(* CODESYS project CodeSys_main_v2.project (continued)
  5ce3da45-db07-42e7-a21c-a00fff4ed8f6|C:\Users\ggb\Documents\#PROJECTS\2016_06_29_Denmark\Visu\CheckBox_1.png
  5ce3da45-db07-42e7-a21c-a00fff4ed8f6|C:\Users\ggb\Documents\#PROJECTS\2016_06_29_Denmark\Visu\Manual_1.png
  5ce3da45-db07-42e7-a21c-a00fff4ed8f6|C:\Users\ggb\Documents\#PROJECTS\2016_06_29_Denmark\Pictures\071-030_Modul Trocknen.jpg
  5ce3da45-db07-42e7-a21c-a00fff4ed8f6|C:\Users\ggb\Documents\#PROJECTS\2016_06_29_Denmark\Visu\English.gif
  5ce3da45-db07-42e7-a21c-a00fff4ed8f6|C:\Users\ggb\Documents\#PROJECTS\2016_06_29_Denmark\Visu\Home_1.png
  5ce3da45-db07-42e7-a21c-a00fff4ed8f6|C:\Users\ggb\Documents\#PROJECTS\2016_06_29_Denmark\Visu\LeftArrow_Bold.png
  5ce3da45-db07-42e7-a21c-a00fff4ed8f6|C:\Users\ggb\Documents\#PROJECTS\2016_06_29_Denmark\Pictures\071-050a_Bohren EA.jpg
  5ce3da45-db07-42e7-a21c-a00fff4ed8f6|C:\Users\ggb\Documents\#PROJECTS\2016_06_29_Denmark\Visu\Parameters_0.png
  Data Types/
    HMI and SCADA/
      data type st_WinCC
      data type st_ManualWorkplace
      CDPX/
        data type st_StopperSensorSignals
        data type st_InterctiveErrors
        data type st_Errors
        data type st_ConveyorSignals
        data type st_AppButtonControl
        data type st_StopperButtonState
        data type st_CdpxButtonState
        data type st_AppSensors
        data type st_ConveyorButtonState
      data type st_ButtonState
      data type st_TransitionData
    SAP/
      sub_structures/
        data type st_Par_Req
        data type st_Start_Req
        data type st_Com
        data type st_Start_Res
        data type st_Comp_Req
        data type st_Comp_Res
      ManualWork/
        data type st_MesRcvData_ManualWork
      data type st_CompleteSfc
      data type st_ParametricData
      data type st_StartSfc
    Error/
      data type st_InteractiveError
      data type st_RobotError
      data type u_Error
      data type st_Error
      data type st_ErrorWords
      data type st_ErrorEvent
    data type st_GetShuntId
    Application/
      data type st_AppControl
      data type st_AppSettings
      data type st_AppState
      data type st_AppInfo
  5ce3da45-db07-42e7-a21c-a00fff4ed8f6|C:\Users\ggb\Documents\#PROJECTS\2016_06_29_Denmark\Visu\Plus.png
  5ce3da45-db07-42e7-a21c-a00fff4ed8f6|C:\Users\ggb\Documents\#PROJECTS\2016_06_29_Denmark\Visu\Settings_1.png
  5ce3da45-db07-42e7-a21c-a00fff4ed8f6|C:\Users\ggb\Documents\#PROJECTS\2016_06_29_Denmark\Visu\Settings_0.png
  5ce3da45-db07-42e7-a21c-a00fff4ed8f6|C:\Users\ggb\Documents\#PROJECTS\2016_06_29_Denmark\Visu\Settings_0.png
  5ce3da45-db07-42e7-a21c-a00fff4ed8f6|C:\Users\ggb\Documents\#PROJECTS\2016_06_29_Denmark\Visu\Parameters_1.png
  5ce3da45-db07-42e7-a21c-a00fff4ed8f6|C:\Users\ggb\Documents\#PROJECTS\2016_06_29_Denmark\Visu\English.gif
  5ce3da45-db07-42e7-a21c-a00fff4ed8f6|C:\Users\ggb\Documents\#PROJECTS\2016_06_29_Denmark\Visu\RightArrow.png
  5ce3da45-db07-42e7-a21c-a00fff4ed8f6|C:\Users\ggb\Documents\#PROJECTS\2016_06_29_Denmark\Pictures\071-050a_Bohren EA.jpg
  5ce3da45-db07-42e7-a21c-a00fff4ed8f6|C:\Users\ggb\Documents\#PROJECTS\2016_06_29_Denmark\Visu\CheckBox_0.png
  5ce3da45-db07-42e7-a21c-a00fff4ed8f6|C:\Users\ggb\Documents\#PROJECTS\2016_06_29_Denmark\Visu\English.gif
  5ce3da45-db07-42e7-a21c-a00fff4ed8f6|C:\Users\ggb\Documents\#PROJECTS\2016_06_29_Denmark\Visu\Stopper.jpg
  5ce3da45-db07-42e7-a21c-a00fff4ed8f6|C:\Users\ggb\Documents\#PROJECTS\2016_06_29_Denmark\Visu\CheckBox_1.png
  5ce3da45-db07-42e7-a21c-a00fff4ed8f6|C:\Users\ggb\Documents\#PROJECTS\2016_06_29_Denmark\Visu\Plus.png
  5ce3da45-db07-42e7-a21c-a00fff4ed8f6|C:\Users\ggb\Documents\#PROJECTS\2016_06_29_Denmark\Pictures\071-046b_Magazin.jpg
  5ce3da45-db07-42e7-a21c-a00fff4ed8f6|C:\Users\ggb\Documents\#PROJECTS\2016_06_29_Denmark\Pictures\cpFactory_Conveyor.png
  5ce3da45-db07-42e7-a21c-a00fff4ed8f6|C:\Users\ggb\Documents\#PROJECTS\2016_06_29_Denmark\Visu\English.gif
  5ce3da45-db07-42e7-a21c-a00fff4ed8f6|C:\Users\ggb\Documents\#PROJECTS\2016_06_29_Denmark\Visu\Parameters_1.png
  5ce3da45-db07-42e7-a21c-a00fff4ed8f6|C:\Users\ggb\Documents\#PROJECTS\2016_06_29_Denmark\Visu\RightArrow.png
  5ce3da45-db07-42e7-a21c-a00fff4ed8f6|C:\Users\ggb\Documents\#PROJECTS\2016_06_29_Denmark\Visu\LeftArrow_Bold.png
  5ce3da45-db07-42e7-a21c-a00fff4ed8f6|C:\Users\ggb\Documents\#PROJECTS\2016_06_29_Denmark\Visu\Manual_1.png
  5ce3da45-db07-42e7-a21c-a00fff4ed8f6|C:\Users\ggb\Documents\#PROJECTS\2016_06_29_Denmark\Visu\Plus.png
  5ce3da45-db07-42e7-a21c-a00fff4ed8f6|C:\Users\ggb\Documents\#PROJECTS\2016_06_29_Denmark\Visu\FESTO.png
  5ce3da45-db07-42e7-a21c-a00fff4ed8f6|C:\Users\ggb\Documents\#PROJECTS\2016_06_29_Denmark\Visu\Parameters_0.png
  5ce3da45-db07-42e7-a21c-a00fff4ed8f6|C:\Users\ggb\Documents\#PROJECTS\2016_06_29_Denmark\Pictures\071-046b_Magazin.jpg
  5ce3da45-db07-42e7-a21c-a00fff4ed8f6|C:\Users\ggb\Documents\#PROJECTS\2016_06_29_Denmark\Visu\LeftArrow_Bold.png
  5ce3da45-db07-42e7-a21c-a00fff4ed8f6|C:\Users\ggb\Documents\#PROJECTS\2016_06_29_Denmark\Visu\Home_0.png
  5ce3da45-db07-42e7-a21c-a00fff4ed8f6|C:\Users\ggb\Documents\#PROJECTS\2016_06_29_Denmark\Visu\Home_1.png
  5ce3da45-db07-42e7-a21c-a00fff4ed8f6|C:\Users\ggb\Documents\#PROJECTS\2016_06_29_Denmark\Visu\German.gif
  5ce3da45-db07-42e7-a21c-a00fff4ed8f6|C:\Users\ggb\Documents\#PROJECTS\2016_06_29_Denmark\Visu\Stopper.jpg
  5ce3da45-db07-42e7-a21c-a00fff4ed8f6|C:\Users\ggb\Documents\#PROJECTS\2016_06_29_Denmark\Visu\RightArrow.png
  5ce3da45-db07-42e7-a21c-a00fff4ed8f6|C:\Users\ggb\Documents\#PROJECTS\2016_06_29_Denmark\Visu\Home_0.png
  5ce3da45-db07-42e7-a21c-a00fff4ed8f6|C:\Users\ggb\Documents\#PROJECTS\2016_06_29_Denmark\Visu\Home_1.png
  5ce3da45-db07-42e7-a21c-a00fff4ed8f6|C:\Users\ggb\Documents\#PROJECTS\2016_06_29_Denmark\Visu\Home_1.png
  5ce3da45-db07-42e7-a21c-a00fff4ed8f6|C:\Users\ggb\Documents\#PROJECTS\2016_06_29_Denmark\Visu\FESTO.png
  5ce3da45-db07-42e7-a21c-a00fff4ed8f6|C:\Users\ggb\Documents\#PROJECTS\2016_06_29_Denmark\Visu\Home_1.png
  5ce3da45-db07-42e7-a21c-a00fff4ed8f6|C:\Users\ggb\Documents\#PROJECTS\2016_06_29_Denmark\Visu\CheckBox_1.png
  5ce3da45-db07-42e7-a21c-a00fff4ed8f6|C:\Users\ggb\Documents\#PROJECTS\2016_06_29_Denmark\Visu\CheckBox_0.png
  5ce3da45-db07-42e7-a21c-a00fff4ed8f6|C:\Users\ggb\Documents\#PROJECTS\2016_06_29_Denmark\Visu\CheckBox_0.png
  5ce3da45-db07-42e7-a21c-a00fff4ed8f6|C:\Users\ggb\Documents\#PROJECTS\2016_06_29_Denmark\Pictures\Cam.jpg
  5ce3da45-db07-42e7-a21c-a00fff4ed8f6|C:\Users\ggb\Documents\#PROJECTS\2016_06_29_Denmark\Visu\Settings_1.png
  5ce3da45-db07-42e7-a21c-a00fff4ed8f6|C:\Users\ggb\Documents\#PROJECTS\2016_06_29_Denmark\Visu\RightArrow_Bold.png
  5ce3da45-db07-42e7-a21c-a00fff4ed8f6|C:\Users\ggb\Documents\#PROJECTS\2016_06_29_Denmark\Visu\RightArrow_Bold.png
  5ce3da45-db07-42e7-a21c-a00fff4ed8f6|C:\Users\ggb\Documents\#PROJECTS\2016_06_29_Denmark\Visu\CheckBox_1.png
  5ce3da45-db07-42e7-a21c-a00fff4ed8f6|C:\Users\ggb\Documents\#PROJECTS\2016_06_29_Denmark\Visu\Settings_0.png
  5ce3da45-db07-42e7-a21c-a00fff4ed8f6|C:\Users\ggb\Documents\#PROJECTS\2016_06_29_Denmark\Visu\Home_0.png
  5ce3da45-db07-42e7-a21c-a00fff4ed8f6|C:\Users\ggb\Documents\#PROJECTS\2016_06_29_Denmark\Pictures\cpFactory_Bypass.png
  5ce3da45-db07-42e7-a21c-a00fff4ed8f6|C:\Users\ggb\Documents\#PROJECTS\2016_06_29_Denmark\Visu\LeftArrow_Bold.png
  5ce3da45-db07-42e7-a21c-a00fff4ed8f6|C:\Users\ggb\Documents\#PROJECTS\2016_06_29_Denmark\Visu\RightArrow.png
  5ce3da45-db07-42e7-a21c-a00fff4ed8f6|C:\Users\ggb\Documents\#PROJECTS\2016_06_29_Denmark\Visu\RightArrow.png
  5ce3da45-db07-42e7-a21c-a00fff4ed8f6|C:\Users\ggb\Documents\#PROJECTS\2016_06_29_Denmark\Visu\RightArrow_Bold.png
  5ce3da45-db07-42e7-a21c-a00fff4ed8f6|C:\Users\ggb\Documents\#PROJECTS\2016_06_29_Denmark\Visu\FESTO.png
  5ce3da45-db07-42e7-a21c-a00fff4ed8f6|C:\Users\ggb\Documents\#PROJECTS\2016_06_29_Denmark\Pictures\cpFactory_Bypass.png
  5ce3da45-db07-42e7-a21c-a00fff4ed8f6|C:\Users\ggb\Documents\#PROJECTS\2016_06_29_Denmark\Visu\Settings_0.png
  5ce3da45-db07-42e7-a21c-a00fff4ed8f6|C:\Users\ggb\Documents\#PROJECTS\2016_06_29_Denmark\Pictures\071-030_Modul Trocknen.jpg
  5ce3da45-db07-42e7-a21c-a00fff4ed8f6|C:\Users\ggb\Documents\#PROJECTS\2016_06_29_Denmark\Visu\RightArrow_Bold.png
  5ce3da45-db07-42e7-a21c-a00fff4ed8f6|C:\Users\ggb\Documents\#PROJECTS\2016_06_29_Denmark\Pictures\071-046b_Magazin.jpg
  5ce3da45-db07-42e7-a21c-a00fff4ed8f6|C:\Users\ggb\Documents\#PROJECTS\2016_06_29_Denmark\Pictures\cpFactory_Bypass.png
  Programs/
    function block TrafficStopper [ST]: _DefaultMode, _ModuleCalls
    function block StopperWithMes [ST]: _MesMode, _DefaultMode, _ModuleCalls, _SapMode
    function block SwitchWithoutMes [ST]: _SapMode, _MesMode, _DefaultMode, _ModuleCalls
    Tools/
      function block ErrorFifo [ST]
      function block MovCntr2B2M [LD]
      function DateFormat [ST]
      function block MovCntr3B3M [LD]
      program ErrorCpyHMI [ST]
      program ErrorCpyWinCC [ST]
    Visu/
      program VisuProgramStp [ST]
    function block SwitchWithMes [ST]: _DefaultMode, _ModuleCalls, _SapMode, _MesMode
  5ce3da45-db07-42e7-a21c-a00fff4ed8f6|C:\Users\ggb\Documents\#PROJECTS\2016_06_29_Denmark\Visu\Home_1.png
  5ce3da45-db07-42e7-a21c-a00fff4ed8f6|C:\Users\ggb\Documents\#PROJECTS\2016_06_29_Denmark\Pictures\cpFactory_Bypass.png
  5ce3da45-db07-42e7-a21c-a00fff4ed8f6|C:\Users\ggb\Documents\#PROJECTS\2016_06_29_Denmark\Visu\CheckBox_0.png
  5ce3da45-db07-42e7-a21c-a00fff4ed8f6|C:\Users\ggb\Documents\#PROJECTS\2016_06_29_Denmark\Pictures\071-046b_Magazin.jpg
  5ce3da45-db07-42e7-a21c-a00fff4ed8f6|C:\Users\ggb\Documents\#PROJECTS\2016_06_29_Denmark\Visu\German.gif
  5ce3da45-db07-42e7-a21c-a00fff4ed8f6|C:\Users\ggb\Documents\#PROJECTS\2016_06_29_Denmark\Visu\RightArrow_Bold.png
  5ce3da45-db07-42e7-a21c-a00fff4ed8f6|C:\Users\ggb\Documents\#PROJECTS\2016_06_29_Denmark\Visu\English.gif
  5ce3da45-db07-42e7-a21c-a00fff4ed8f6|C:\Users\ggb\Documents\#PROJECTS\2016_06_29_Denmark\Pictures\Kuka_Agilus.png
  5ce3da45-db07-42e7-a21c-a00fff4ed8f6|C:\Users\ggb\Documents\#PROJECTS\2016_06_29_Denmark\Visu\Parameters_1.png
  5ce3da45-db07-42e7-a21c-a00fff4ed8f6|C:\Users\ggb\Documents\#PROJECTS\2016_06_29_Denmark\Visu\FESTO.png
  5ce3da45-db07-42e7-a21c-a00fff4ed8f6|C:\Users\ggb\Documents\#PROJECTS\2016_06_29_Denmark\Pictures\071-046b_Magazin.jpg
  5ce3da45-db07-42e7-a21c-a00fff4ed8f6|C:\Users\ggb\Documents\#PROJECTS\2016_06_29_Denmark\Visu\German.gif
  5ce3da45-db07-42e7-a21c-a00fff4ed8f6|C:\Users\ggb\Documents\#PROJECTS\2016_06_29_Denmark\Visu\Settings_0.png
  5ce3da45-db07-42e7-a21c-a00fff4ed8f6|C:\Users\ggb\Documents\#PROJECTS\2016_06_29_Denmark\Visu\Plus.png
  5ce3da45-db07-42e7-a21c-a00fff4ed8f6|C:\Users\ggb\Documents\#PROJECTS\2016_06_29_Denmark\Visu\Settings_1.png
  5ce3da45-db07-42e7-a21c-a00fff4ed8f6|C:\Users\ggb\Documents\#PROJECTS\2016_06_29_Denmark\Visu\Settings_0.png
  5ce3da45-db07-42e7-a21c-a00fff4ed8f6|C:\Users\ggb\Documents\#PROJECTS\2016_06_29_Denmark\Visu\CheckBox_1.png
  5ce3da45-db07-42e7-a21c-a00fff4ed8f6|C:\Users\ggb\Documents\#PROJECTS\2016_06_29_Denmark\Visu\German.gif
  5ce3da45-db07-42e7-a21c-a00fff4ed8f6|C:\Users\ggb\Documents\#PROJECTS\2016_06_29_Denmark\Visu\Plus.png
  5ce3da45-db07-42e7-a21c-a00fff4ed8f6|C:\Users\ggb\Documents\#PROJECTS\2016_06_29_Denmark\Pictures\071-060_Kameraprüfen.jpg
  5ce3da45-db07-42e7-a21c-a00fff4ed8f6|C:\Users\ggb\Documents\#PROJECTS\2016_06_29_Denmark\Visu\Manual_0.png
  5ce3da45-db07-42e7-a21c-a00fff4ed8f6|C:\Users\ggb\Documents\#PROJECTS\2016_06_29_Denmark\Visu\Settings_1.png
  5ce3da45-db07-42e7-a21c-a00fff4ed8f6|C:\Users\ggb\Documents\#PROJECTS\2016_06_29_Denmark\Pictures\071-050a_Bohren EA.jpg
  5ce3da45-db07-42e7-a21c-a00fff4ed8f6|C:\Users\ggb\Documents\#PROJECTS\2016_06_29_Denmark\Visu\Settings_1.png
  5ce3da45-db07-42e7-a21c-a00fff4ed8f6|C:\Users\ggb\Documents\#PROJECTS\2016_06_29_Denmark\Pictures\071-030_Modul Trocknen.jpg
  5ce3da45-db07-42e7-a21c-a00fff4ed8f6|C:\Users\ggb\Documents\#PROJECTS\2016_06_29_Denmark\Visu\LeftArrow_Bold.png
  5ce3da45-db07-42e7-a21c-a00fff4ed8f6|C:\Users\ggb\Documents\#PROJECTS\2016_06_29_Denmark\Pictures\071-030_Modul Trocknen.jpg
  5ce3da45-db07-42e7-a21c-a00fff4ed8f6|C:\Users\ggb\Documents\#PROJECTS\2016_06_29_Denmark\Pictures\071-046b_Magazin.jpg
  5ce3da45-db07-42e7-a21c-a00fff4ed8f6|C:\Users\ggb\Documents\#PROJECTS\2016_06_29_Denmark\Pictures\cpFactory_Bypass.png
  5ce3da45-db07-42e7-a21c-a00fff4ed8f6|C:\Users\ggb\Documents\#PROJECTS\2016_06_29_Denmark\Visu\Plus.png
  5ce3da45-db07-42e7-a21c-a00fff4ed8f6|C:\Users\ggb\Documents\#PROJECTS\2016_06_29_Denmark\Visu\FESTO.png
  5ce3da45-db07-42e7-a21c-a00fff4ed8f6|C:\Users\ggb\Documents\#PROJECTS\2016_06_29_Denmark\Visu\English.gif
  5ce3da45-db07-42e7-a21c-a00fff4ed8f6|C:\Users\ggb\Documents\#PROJECTS\2016_06_29_Denmark\Visu\Stopper.jpg
  5ce3da45-db07-42e7-a21c-a00fff4ed8f6|C:\Users\ggb\Documents\#PROJECTS\2016_06_29_Denmark\Visu\Stopper.jpg
  5ce3da45-db07-42e7-a21c-a00fff4ed8f6|C:\Users\ggb\Documents\#PROJECTS\2016_06_29_Denmark\Pictures\071-030_Modul Trocknen.jpg
  5ce3da45-db07-42e7-a21c-a00fff4ed8f6|C:\Users\ggb\Documents\#PROJECTS\2016_06_29_Denmark\Pictures\cpFactory_Bypass.png
  5ce3da45-db07-42e7-a21c-a00fff4ed8f6|C:\Users\ggb\Documents\#PROJECTS\2016_06_29_Denmark\Visu\CheckBox_0.png
  5ce3da45-db07-42e7-a21c-a00fff4ed8f6|C:\Users\ggb\Documents\#PROJECTS\2016_06_29_Denmark\Visu\CheckBox_0.png
  5ce3da45-db07-42e7-a21c-a00fff4ed8f6|C:\Users\ggb\Documents\#PROJECTS\2016_06_29_Denmark\Visu\Stopper.jpg
  5ce3da45-db07-42e7-a21c-a00fff4ed8f6|C:\Users\ggb\Documents\#PROJECTS\2016_06_29_Denmark\Pictures\cpFactory_Conveyor.png
  5ce3da45-db07-42e7-a21c-a00fff4ed8f6|C:\Users\ggb\Documents\#PROJECTS\2016_06_29_Denmark\Visu\Settings_0.png
  5ce3da45-db07-42e7-a21c-a00fff4ed8f6|C:\Users\ggb\Documents\#PROJECTS\2016_06_29_Denmark\Visu\Parameters_0.png
  5ce3da45-db07-42e7-a21c-a00fff4ed8f6|C:\Users\ggb\Documents\#PROJECTS\2016_06_29_Denmark\Visu\Home_1.png
  5ce3da45-db07-42e7-a21c-a00fff4ed8f6|C:\Users\ggb\Documents\#PROJECTS\2016_06_29_Denmark\Pictures\071-050a_Bohren EA.jpg
  5ce3da45-db07-42e7-a21c-a00fff4ed8f6|C:\Users\ggb\Documents\#PROJECTS\2016_06_29_Denmark\Visu\Manual_1.png
  5ce3da45-db07-42e7-a21c-a00fff4ed8f6|C:\Users\ggb\Documents\#PROJECTS\2016_06_29_Denmark\Visu\Stopper.jpg
  5ce3da45-db07-42e7-a21c-a00fff4ed8f6|C:\Users\ggb\Documents\#PROJECTS\2016_06_29_Denmark\Pictures\071-030_Modul Trocknen.jpg
  5ce3da45-db07-42e7-a21c-a00fff4ed8f6|C:\Users\ggb\Documents\#PROJECTS\2016_06_29_Denmark\Visu\CheckBox_0.png
  5ce3da45-db07-42e7-a21c-a00fff4ed8f6|C:\Users\ggb\Documents\#PROJECTS\2016_06_29_Denmark\Visu\CheckBox_1.png
  5ce3da45-db07-42e7-a21c-a00fff4ed8f6|C:\Users\ggb\Documents\#PROJECTS\2016_06_29_Denmark\Visu\LeftArrow_Bold.png
  5ce3da45-db07-42e7-a21c-a00fff4ed8f6|C:\Users\ggb\Documents\#PROJECTS\2016_06_29_Denmark\Pictures\cpFactory_Bypass.png
  5ce3da45-db07-42e7-a21c-a00fff4ed8f6|C:\Users\ggb\Documents\#PROJECTS\2016_06_29_Denmark\Visu\LeftArrow_Bold.png
  Global Variables/
    global variables fromCDPX
    global variables Standards
    global variables toCDPX
    global variables SAP
    global variables SAPInit
    global variables SAPHMI
  5ce3da45-db07-42e7-a21c-a00fff4ed8f6|C:\Users\ggb\Documents\#PROJECTS\2016_06_29_Denmark\Visu\CheckBox_0.png
  5ce3da45-db07-42e7-a21c-a00fff4ed8f6|C:\Users\ggb\Documents\#PROJECTS\2016_06_29_Denmark\Pictures\cpFactory_Conveyor.png
  5ce3da45-db07-42e7-a21c-a00fff4ed8f6|C:\Users\ggb\Documents\#PROJECTS\2016_06_29_Denmark\Pictures\071-046b_Magazin.jpg
  5ce3da45-db07-42e7-a21c-a00fff4ed8f6|C:\Users\ggb\Documents\#PROJECTS\2016_06_29_Denmark\Visu\RightArrow.png
  5ce3da45-db07-42e7-a21c-a00fff4ed8f6|C:\Users\ggb\Documents\#PROJECTS\2016_06_29_Denmark\Pictures\cpFactory_Bypass.png
  5ce3da45-db07-42e7-a21c-a00fff4ed8f6|C:\Users\ggb\Documents\#PROJECTS\2016_06_29_Denmark\Pictures\071-060_Kameraprüfen.jpg
  5ce3da45-db07-42e7-a21c-a00fff4ed8f6|C:\Users\ggb\Documents\#PROJECTS\2016_06_29_Denmark\Visu\German.gif
  5ce3da45-db07-42e7-a21c-a00fff4ed8f6|C:\Users\ggb\Documents\#PROJECTS\2016_06_29_Denmark\Visu\CheckBox_0.png
  5ce3da45-db07-42e7-a21c-a00fff4ed8f6|C:\Users\ggb\Documents\#PROJECTS\2016_06_29_Denmark\Visu\Settings_0.png
  5ce3da45-db07-42e7-a21c-a00fff4ed8f6|C:\Users\ggb\Documents\#PROJECTS\2016_06_29_Denmark\Visu\CheckBox_1.png
  5ce3da45-db07-42e7-a21c-a00fff4ed8f6|C:\Users\ggb\Documents\#PROJECTS\2016_06_29_Denmark\Visu\FESTO.png
  5ce3da45-db07-42e7-a21c-a00fff4ed8f6|C:\Users\ggb\Documents\#PROJECTS\2016_06_29_Denmark\Visu\CheckBox_0.png
  5ce3da45-db07-42e7-a21c-a00fff4ed8f6|C:\Users\ggb\Documents\#PROJECTS\2016_06_29_Denmark\Pictures\cpFactory_Conveyor.png
  5ce3da45-db07-42e7-a21c-a00fff4ed8f6|C:\Users\ggb\Documents\#PROJECTS\2016_06_29_Denmark\Visu\CheckBox_1.png
  5ce3da45-db07-42e7-a21c-a00fff4ed8f6|C:\Users\ggb\Documents\#PROJECTS\2016_06_29_Denmark\Pictures\cpFactory_Conveyor.png
  5ce3da45-db07-42e7-a21c-a00fff4ed8f6|C:\Users\ggb\Documents\#PROJECTS\2016_06_29_Denmark\Pictures\071-050a_Bohren EA.jpg
  5ce3da45-db07-42e7-a21c-a00fff4ed8f6|C:\Users\ggb\Documents\#PROJECTS\2016_06_29_Denmark\Visu\Parameters_0.png
  5ce3da45-db07-42e7-a21c-a00fff4ed8f6|C:\Users\ggb\Documents\#PROJECTS\2016_06_29_Denmark\Visu\CheckBox_1.png
  5ce3da45-db07-42e7-a21c-a00fff4ed8f6|C:\Users\ggb\Documents\#PROJECTS\2016_06_29_Denmark\Visu\Home_1.png
  5ce3da45-db07-42e7-a21c-a00fff4ed8f6|C:\Users\ggb\Documents\#PROJECTS\2016_06_29_Denmark\Pictures\071-060_Kameraprüfen.jpg
  5ce3da45-db07-42e7-a21c-a00fff4ed8f6|C:\Users\ggb\Documents\#PROJECTS\2016_06_29_Denmark\Visu\English.gif
  5ce3da45-db07-42e7-a21c-a00fff4ed8f6|C:\Users\ggb\Documents\#PROJECTS\2016_06_29_Denmark\Pictures\cpFactory_Bypass.png
  5ce3da45-db07-42e7-a21c-a00fff4ed8f6|C:\Users\ggb\Documents\#PROJECTS\2016_06_29_Denmark\Visu\Parameters_1.png
  5ce3da45-db07-42e7-a21c-a00fff4ed8f6|C:\Users\ggb\Documents\#PROJECTS\2016_06_29_Denmark\Visu\Manual_1.png
  5ce3da45-db07-42e7-a21c-a00fff4ed8f6|C:\Users\ggb\Documents\#PROJECTS\2016_06_29_Denmark\Visu\CheckBox_0.png
  5ce3da45-db07-42e7-a21c-a00fff4ed8f6|C:\Users\ggb\Documents\#PROJECTS\2016_06_29_Denmark\Visu\Manual_0.png
  5ce3da45-db07-42e7-a21c-a00fff4ed8f6|C:\Users\ggb\Documents\#PROJECTS\2016_06_29_Denmark\Visu\Manual_0.png
  5ce3da45-db07-42e7-a21c-a00fff4ed8f6|C:\Users\ggb\Documents\#PROJECTS\2016_06_29_Denmark\Visu\Home_1.png
  5ce3da45-db07-42e7-a21c-a00fff4ed8f6|C:\Users\ggb\Documents\#PROJECTS\2016_06_29_Denmark\Pictures\071-046b_Magazin.jpg
  5ce3da45-db07-42e7-a21c-a00fff4ed8f6|C:\Users\ggb\Documents\#PROJECTS\2016_06_29_Denmark\Visu\English.gif
  5ce3da45-db07-42e7-a21c-a00fff4ed8f6|C:\Users\ggb\Documents\#PROJECTS\2016_06_29_Denmark\Pictures\cpFactory_Conveyor.png
  5ce3da45-db07-42e7-a21c-a00fff4ed8f6|C:\Users\ggb\Documents\#PROJECTS\2016_06_29_Denmark\Pictures\071-050a_Bohren EA.jpg
  5ce3da45-db07-42e7-a21c-a00fff4ed8f6|C:\Users\ggb\Documents\#PROJECTS\2016_06_29_Denmark\Visu\English.gif
  5ce3da45-db07-42e7-a21c-a00fff4ed8f6|C:\Users\ggb\Documents\#PROJECTS\2016_06_29_Denmark\Visu\Parameters_1.png
  5ce3da45-db07-42e7-a21c-a00fff4ed8f6|C:\Users\ggb\Documents\#PROJECTS\2016_06_29_Denmark\Visu\RightArrow_Bold.png
  5ce3da45-db07-42e7-a21c-a00fff4ed8f6|C:\Users\ggb\Documents\#PROJECTS\2016_06_29_Denmark\Visu\FESTO.png
  5ce3da45-db07-42e7-a21c-a00fff4ed8f6|C:\Users\ggb\Documents\#PROJECTS\2016_06_29_Denmark\Pictures\071-050a_Bohren EA.jpg
  5ce3da45-db07-42e7-a21c-a00fff4ed8f6|C:\Users\ggb\Documents\#PROJECTS\2016_06_29_Denmark\Pictures\071-046b_Magazin.jpg
  5ce3da45-db07-42e7-a21c-a00fff4ed8f6|C:\Users\ggb\Documents\#PROJECTS\2016_06_29_Denmark\Visu\RightArrow_Bold.png
  5ce3da45-db07-42e7-a21c-a00fff4ed8f6|C:\Users\ggb\Documents\#PROJECTS\2016_06_29_Denmark\Visu\Parameters_0.png
  5ce3da45-db07-42e7-a21c-a00fff4ed8f6|C:\Users\ggb\Documents\#PROJECTS\2016_06_29_Denmark\Pictures\cpFactory_Conveyor.png
  5ce3da45-db07-42e7-a21c-a00fff4ed8f6|C:\Users\ggb\Documents\#PROJECTS\2016_06_29_Denmark\Visu\Home_0.png
  5ce3da45-db07-42e7-a21c-a00fff4ed8f6|C:\Users\ggb\Documents\#PROJECTS\2016_06_29_Denmark\Visu\LeftArrow_Bold.png
  5ce3da45-db07-42e7-a21c-a00fff4ed8f6|C:\Users\ggb\Documents\#PROJECTS\2016_06_29_Denmark\Visu\Parameters_0.png
  5ce3da45-db07-42e7-a21c-a00fff4ed8f6|C:\Users\ggb\Documents\#PROJECTS\2016_06_29_Denmark\Visu\Manual_0.png
  5ce3da45-db07-42e7-a21c-a00fff4ed8f6|C:\Users\ggb\Documents\#PROJECTS\2016_06_29_Denmark\Visu\Manual_0.png
  5ce3da45-db07-42e7-a21c-a00fff4ed8f6|C:\Users\ggb\Documents\#PROJECTS\2016_06_29_Denmark\Visu\Settings_1.png
  5ce3da45-db07-42e7-a21c-a00fff4ed8f6|C:\Users\ggb\Documents\#PROJECTS\2016_06_29_Denmark\Visu\Home_0.png
  5ce3da45-db07-42e7-a21c-a00fff4ed8f6|C:\Users\ggb\Documents\#PROJECTS\2016_06_29_Denmark\Visu\FESTO.png
  5ce3da45-db07-42e7-a21c-a00fff4ed8f6|C:\Users\ggb\Documents\#PROJECTS\2016_06_29_Denmark\Visu\German.gif
  5ce3da45-db07-42e7-a21c-a00fff4ed8f6|C:\Users\ggb\Documents\#PROJECTS\2016_06_29_Denmark\Visu\Settings_0.png
  5ce3da45-db07-42e7-a21c-a00fff4ed8f6|C:\Users\ggb\Documents\#PROJECTS\2016_06_29_Denmark\Visu\RightArrow_Bold.png
  5ce3da45-db07-42e7-a21c-a00fff4ed8f6|C:\Users\ggb\Documents\#PROJECTS\2016_06_29_Denmark\Visu\Stopper.jpg
  5ce3da45-db07-42e7-a21c-a00fff4ed8f6|C:\Users\ggb\Documents\#PROJECTS\2016_06_29_Denmark\Visu\Parameters_1.png
  5ce3da45-db07-42e7-a21c-a00fff4ed8f6|C:\Users\ggb\Documents\#PROJECTS\2016_06_29_Denmark\Visu\FESTO.png
  5ce3da45-db07-42e7-a21c-a00fff4ed8f6|C:\Users\ggb\Documents\#PROJECTS\2016_06_29_Denmark\Visu\German.gif
  5ce3da45-db07-42e7-a21c-a00fff4ed8f6|C:\Users\ggb\Documents\#PROJECTS\2016_06_29_Denmark\Visu\Home_0.png
  text list GlobalTextList
  5ce3da45-db07-42e7-a21c-a00fff4ed8f6|C:\Users\ggb\Documents\#PROJECTS\2016_06_29_Denmark\Visu\FESTO.png
  5ce3da45-db07-42e7-a21c-a00fff4ed8f6|C:\Users\ggb\Documents\#PROJECTS\2016_06_29_Denmark\Visu\Home_1.png
  5ce3da45-db07-42e7-a21c-a00fff4ed8f6|C:\Users\ggb\Documents\#PROJECTS\2016_06_29_Denmark\Visu\Manual_0.png
  5ce3da45-db07-42e7-a21c-a00fff4ed8f6|C:\Users\ggb\Documents\#PROJECTS\2016_06_29_Denmark\Visu\Stopper.jpg
  5ce3da45-db07-42e7-a21c-a00fff4ed8f6|C:\Users\ggb\Documents\#PROJECTS\2016_06_29_Denmark\Visu\LeftArrow_Bold.png
  5ce3da45-db07-42e7-a21c-a00fff4ed8f6|C:\Users\ggb\Documents\#PROJECTS\2016_06_29_Denmark\Visu\Manual_0.png
  5ce3da45-db07-42e7-a21c-a00fff4ed8f6|C:\Users\ggb\Documents\#PROJECTS\2016_06_29_Denmark\Visu\CheckBox_0.png
  5ce3da45-db07-42e7-a21c-a00fff4ed8f6|C:\Users\ggb\Documents\#PROJECTS\2016_06_29_Denmark\Visu\Plus.png
  5ce3da45-db07-42e7-a21c-a00fff4ed8f6|C:\Users\ggb\Documents\#PROJECTS\2016_06_29_Denmark\Pictures\071-030_Modul Trocknen.jpg
  5ce3da45-db07-42e7-a21c-a00fff4ed8f6|C:\Users\ggb\Documents\#PROJECTS\2016_06_29_Denmark\Visu\Parameters_1.png
  5ce3da45-db07-42e7-a21c-a00fff4ed8f6|C:\Users\ggb\Documents\#PROJECTS\2016_06_29_Denmark\Visu\LeftArrow_Bold.png
  5ce3da45-db07-42e7-a21c-a00fff4ed8f6|C:\Users\ggb\Documents\#PROJECTS\2016_06_29_Denmark\Pictures\cpFactory_Conveyor.png
  5ce3da45-db07-42e7-a21c-a00fff4ed8f6|C:\Users\ggb\Documents\#PROJECTS\2016_06_29_Denmark\Visu\Manual_0.png
  5ce3da45-db07-42e7-a21c-a00fff4ed8f6|C:\Users\ggb\Documents\#PROJECTS\2016_06_29_Denmark\Visu\RightArrow_Bold.png
  5ce3da45-db07-42e7-a21c-a00fff4ed8f6|C:\Users\ggb\Documents\#PROJECTS\2016_06_29_Denmark\Visu\CheckBox_1.png
  5ce3da45-db07-42e7-a21c-a00fff4ed8f6|C:\Users\ggb\Documents\#PROJECTS\2016_06_29_Denmark\Visu\English.gif
  5ce3da45-db07-42e7-a21c-a00fff4ed8f6|C:\Users\ggb\Documents\#PROJECTS\2016_06_29_Denmark\Visu\FESTO.png
  5ce3da45-db07-42e7-a21c-a00fff4ed8f6|C:\Users\ggb\Documents\#PROJECTS\2016_06_29_Denmark\Visu\English.gif
  5ce3da45-db07-42e7-a21c-a00fff4ed8f6|C:\Users\ggb\Documents\#PROJECTS\2016_06_29_Denmark\Pictures\cpFactory_Conveyor.png
  5ce3da45-db07-42e7-a21c-a00fff4ed8f6|C:\Users\ggb\Documents\#PROJECTS\2016_06_29_Denmark\Visu\Parameters_0.png
  5ce3da45-db07-42e7-a21c-a00fff4ed8f6|C:\Users\ggb\Documents\#PROJECTS\2016_06_29_Denmark\Pictures\071-060_Kameraprüfen.jpg
  5ce3da45-db07-42e7-a21c-a00fff4ed8f6|C:\Users\ggb\Documents\#PROJECTS\2016_06_29_Denmark\Pictures\Kuka_Agilus.png
  5ce3da45-db07-42e7-a21c-a00fff4ed8f6|C:\Users\ggb\Documents\#PROJECTS\2016_06_29_Denmark\Pictures\071-046b_Magazin.jpg
  5ce3da45-db07-42e7-a21c-a00fff4ed8f6|C:\Users\ggb\Documents\#PROJECTS\2016_06_29_Denmark\Pictures\cpFactory_Bypass.png
  5ce3da45-db07-42e7-a21c-a00fff4ed8f6|C:\Users\ggb\Documents\#PROJECTS\2016_06_29_Denmark\Visu\LeftArrow_Bold.png
  5ce3da45-db07-42e7-a21c-a00fff4ed8f6|C:\Users\ggb\Documents\#PROJECTS\2016_06_29_Denmark\Pictures\071-030_Modul Trocknen.jpg
  5ce3da45-db07-42e7-a21c-a00fff4ed8f6|C:\Users\ggb\Documents\#PROJECTS\2016_06_29_Denmark\Visu\German.gif
  5ce3da45-db07-42e7-a21c-a00fff4ed8f6|C:\Users\ggb\Documents\#PROJECTS\2016_06_29_Denmark\Visu\Manual_0.png
  5ce3da45-db07-42e7-a21c-a00fff4ed8f6|C:\Users\ggb\Documents\#PROJECTS\2016_06_29_Denmark\Visu\German.gif
  5ce3da45-db07-42e7-a21c-a00fff4ed8f6|C:\Users\ggb\Documents\#PROJECTS\2016_06_29_Denmark\Visu\CheckBox_1.png
  5ce3da45-db07-42e7-a21c-a00fff4ed8f6|C:\Users\ggb\Documents\#PROJECTS\2016_06_29_Denmark\Visu\Home_0.png
  5ce3da45-db07-42e7-a21c-a00fff4ed8f6|C:\Users\ggb\Documents\#PROJECTS\2016_06_29_Denmark\Visu\Settings_1.png
  5ce3da45-db07-42e7-a21c-a00fff4ed8f6|C:\Users\ggb\Documents\#PROJECTS\2016_06_29_Denmark\Visu\Settings_1.png
  5ce3da45-db07-42e7-a21c-a00fff4ed8f6|C:\Users\ggb\Documents\#PROJECTS\2016_06_29_Denmark\Pictures\071-060_Kameraprüfen.jpg
  5ce3da45-db07-42e7-a21c-a00fff4ed8f6|C:\Users\ggb\Documents\#PROJECTS\2016_06_29_Denmark\Visu\FESTO.png
  5ce3da45-db07-42e7-a21c-a00fff4ed8f6|C:\Users\ggb\Documents\#PROJECTS\2016_06_29_Denmark\Visu\Manual_1.png
  5ce3da45-db07-42e7-a21c-a00fff4ed8f6|C:\Users\ggb\Documents\#PROJECTS\2016_06_29_Denmark\Visu\Home_0.png
  5ce3da45-db07-42e7-a21c-a00fff4ed8f6|C:\Users\ggb\Documents\#PROJECTS\2016_06_29_Denmark\Visu\Plus.png
  5ce3da45-db07-42e7-a21c-a00fff4ed8f6|C:\Users\ggb\Documents\#PROJECTS\2016_06_29_Denmark\Pictures\071-030_Modul Trocknen.jpg
  5ce3da45-db07-42e7-a21c-a00fff4ed8f6|C:\Users\ggb\Documents\#PROJECTS\2016_06_29_Denmark\Visu\CheckBox_1.png
  5ce3da45-db07-42e7-a21c-a00fff4ed8f6|C:\Users\ggb\Documents\#PROJECTS\2016_06_29_Denmark\Visu\Stopper.jpg
  5ce3da45-db07-42e7-a21c-a00fff4ed8f6|C:\Users\ggb\Documents\#PROJECTS\2016_06_29_Denmark\Visu\Manual_1.png
  5ce3da45-db07-42e7-a21c-a00fff4ed8f6|C:\Users\ggb\Documents\#PROJECTS\2016_06_29_Denmark\Visu\Manual_0.png
  5ce3da45-db07-42e7-a21c-a00fff4ed8f6|C:\Users\ggb\Documents\#PROJECTS\2016_06_29_Denmark\Visu\FESTO.png
  5ce3da45-db07-42e7-a21c-a00fff4ed8f6|C:\Users\ggb\Documents\#PROJECTS\2016_06_29_Denmark\Visu\Settings_0.png
  5ce3da45-db07-42e7-a21c-a00fff4ed8f6|C:\Users\ggb\Documents\#PROJECTS\2016_06_29_Denmark\Pictures\071-060_Kameraprüfen.jpg
  5ce3da45-db07-42e7-a21c-a00fff4ed8f6|C:\Users\ggb\Documents\#PROJECTS\2016_06_29_Denmark\Visu\Parameters_1.png
  5ce3da45-db07-42e7-a21c-a00fff4ed8f6|C:\Users\ggb\Documents\#PROJECTS\2016_06_29_Denmark\Visu\Settings_0.png
  5ce3da45-db07-42e7-a21c-a00fff4ed8f6|C:\Users\ggb\Documents\#PROJECTS\2016_06_29_Denmark\Pictures\071-046b_Magazin.jpg
  5ce3da45-db07-42e7-a21c-a00fff4ed8f6|C:\Users\ggb\Documents\#PROJECTS\2016_06_29_Denmark\Visu\CheckBox_0.png
  5ce3da45-db07-42e7-a21c-a00fff4ed8f6|C:\Users\ggb\Documents\#PROJECTS\2016_06_29_Denmark\Visu\LeftArrow_Bold.png
  5ce3da45-db07-42e7-a21c-a00fff4ed8f6|C:\Users\ggb\Documents\#PROJECTS\2016_06_29_Denmark\Pictures\071-060_Kameraprüfen.jpg
  5ce3da45-db07-42e7-a21c-a00fff4ed8f6|C:\Users\ggb\Documents\#PROJECTS\2016_06_29_Denmark\Pictures\071-046b_Magazin.jpg
  5ce3da45-db07-42e7-a21c-a00fff4ed8f6|C:\Users\ggb\Documents\#PROJECTS\2016_06_29_Denmark\Visu\Parameters_0.png
  5ce3da45-db07-42e7-a21c-a00fff4ed8f6|C:\Users\ggb\Documents\#PROJECTS\2016_06_29_Denmark\Visu\CheckBox_1.png
  5ce3da45-db07-42e7-a21c-a00fff4ed8f6|C:\Users\ggb\Documents\#PROJECTS\2016_06_29_Denmark\Visu\RightArrow.png
  5ce3da45-db07-42e7-a21c-a00fff4ed8f6|C:\Users\ggb\Documents\#PROJECTS\2016_06_29_Denmark\Visu\FESTO.png
  5ce3da45-db07-42e7-a21c-a00fff4ed8f6|C:\Users\ggb\Documents\#PROJECTS\2016_06_29_Denmark\Visu\LeftArrow_Bold.png
  5ce3da45-db07-42e7-a21c-a00fff4ed8f6|C:\Users\ggb\Documents\#PROJECTS\2016_06_29_Denmark\Visu\Manual_1.png
  5ce3da45-db07-42e7-a21c-a00fff4ed8f6|C:\Users\ggb\Documents\#PROJECTS\2016_06_29_Denmark\Visu\LeftArrow_Bold.png
  5ce3da45-db07-42e7-a21c-a00fff4ed8f6|C:\Users\ggb\Documents\#PROJECTS\2016_06_29_Denmark\Pictures\071-046b_Magazin.jpg
  5ce3da45-db07-42e7-a21c-a00fff4ed8f6|C:\Users\ggb\Documents\#PROJECTS\2016_06_29_Denmark\Visu\RightArrow.png
  5ce3da45-db07-42e7-a21c-a00fff4ed8f6|C:\Users\ggb\Documents\#PROJECTS\2016_06_29_Denmark\Visu\Parameters_0.png
  5ce3da45-db07-42e7-a21c-a00fff4ed8f6|C:\Users\ggb\Documents\#PROJECTS\2016_06_29_Denmark\Visu\Home_0.png
  5ce3da45-db07-42e7-a21c-a00fff4ed8f6|C:\Users\ggb\Documents\#PROJECTS\2016_06_29_Denmark\Visu\Home_0.png
  5ce3da45-db07-42e7-a21c-a00fff4ed8f6|C:\Users\ggb\Documents\#PROJECTS\2016_06_29_Denmark\Visu\Manual_1.png
  5ce3da45-db07-42e7-a21c-a00fff4ed8f6|C:\Users\ggb\Documents\#PROJECTS\2016_06_29_Denmark\Visu\Manual_1.png
  5ce3da45-db07-42e7-a21c-a00fff4ed8f6|C:\Users\ggb\Documents\#PROJECTS\2016_06_29_Denmark\Visu\RightArrow_Bold.png
  5ce3da45-db07-42e7-a21c-a00fff4ed8f6|C:\Users\ggb\Documents\#PROJECTS\2016_06_29_Denmark\Visu\Home_0.png
  5ce3da45-db07-42e7-a21c-a00fff4ed8f6|C:\Users\ggb\Documents\#PROJECTS\2016_06_29_Denmark\Visu\German.gif
  5ce3da45-db07-42e7-a21c-a00fff4ed8f6|C:\Users\ggb\Documents\#PROJECTS\2016_06_29_Denmark\Pictures\071-060_Kameraprüfen.jpg
  5ce3da45-db07-42e7-a21c-a00fff4ed8f6|C:\Users\ggb\Documents\#PROJECTS\2016_06_29_Denmark\Pictures\071-030_Modul Trocknen.jpg
  5ce3da45-db07-42e7-a21c-a00fff4ed8f6|C:\Users\ggb\Documents\#PROJECTS\2016_06_29_Denmark\Visu\Home_0.png
  5ce3da45-db07-42e7-a21c-a00fff4ed8f6|C:\Users\ggb\Documents\#PROJECTS\2016_06_29_Denmark\Visu\Settings_1.png
  5ce3da45-db07-42e7-a21c-a00fff4ed8f6|C:\Users\ggb\Documents\#PROJECTS\2016_06_29_Denmark\Pictures\071-060_Kameraprüfen.jpg
  5ce3da45-db07-42e7-a21c-a00fff4ed8f6|C:\Users\ggb\Documents\#PROJECTS\2016_06_29_Denmark\Visu\Settings_1.png
  5ce3da45-db07-42e7-a21c-a00fff4ed8f6|C:\Users\ggb\Documents\#PROJECTS\2016_06_29_Denmark\Visu\Stopper.jpg
  5ce3da45-db07-42e7-a21c-a00fff4ed8f6|C:\Users\ggb\Documents\#PROJECTS\2016_06_29_Denmark\Visu\Manual_1.png
  5ce3da45-db07-42e7-a21c-a00fff4ed8f6|C:\Users\ggb\Documents\#PROJECTS\2016_06_29_Denmark\Pictures\cpFactory_Bypass.png
  5ce3da45-db07-42e7-a21c-a00fff4ed8f6|C:\Users\ggb\Documents\#PROJECTS\2016_06_29_Denmark\Visu\CheckBox_1.png
  5ce3da45-db07-42e7-a21c-a00fff4ed8f6|C:\Users\ggb\Documents\#PROJECTS\2016_06_29_Denmark\Pictures\cpFactory_Conveyor.png
  5ce3da45-db07-42e7-a21c-a00fff4ed8f6|C:\Users\ggb\Documents\#PROJECTS\2016_06_29_Denmark\Visu\Home_1.png
  5ce3da45-db07-42e7-a21c-a00fff4ed8f6|C:\Users\ggb\Documents\#PROJECTS\2016_06_29_Denmark\Visu\Home_1.png
  5ce3da45-db07-42e7-a21c-a00fff4ed8f6|C:\Users\ggb\Documents\#PROJECTS\2016_06_29_Denmark\Visu\RightArrow_Bold.png
  5ce3da45-db07-42e7-a21c-a00fff4ed8f6|C:\Users\ggb\Documents\#PROJECTS\2016_06_29_Denmark\Visu\RightArrow_Bold.png
  5ce3da45-db07-42e7-a21c-a00fff4ed8f6|C:\Users\ggb\Documents\#PROJECTS\2016_06_29_Denmark\Visu\Settings_0.png
  5ce3da45-db07-42e7-a21c-a00fff4ed8f6|C:\Users\ggb\Documents\#PROJECTS\2016_06_29_Denmark\Visu\English.gif
  5ce3da45-db07-42e7-a21c-a00fff4ed8f6|C:\Users\ggb\Documents\#PROJECTS\2016_06_29_Denmark\Pictures\071-060_Kameraprüfen.jpg
  5ce3da45-db07-42e7-a21c-a00fff4ed8f6|C:\Users\ggb\Documents\#PROJECTS\2016_06_29_Denmark\Visu\Parameters_1.png
  5ce3da45-db07-42e7-a21c-a00fff4ed8f6|C:\Users\ggb\Documents\#PROJECTS\2016_06_29_Denmark\Visu\Plus.png
  5ce3da45-db07-42e7-a21c-a00fff4ed8f6|C:\Users\ggb\Documents\#PROJECTS\2016_06_29_Denmark\Visu\Stopper.jpg
  5ce3da45-db07-42e7-a21c-a00fff4ed8f6|C:\Users\ggb\Documents\#PROJECTS\2016_06_29_Denmark\Visu\Parameters_1.png
  5ce3da45-db07-42e7-a21c-a00fff4ed8f6|C:\Users\ggb\Documents\#PROJECTS\2016_06_29_Denmark\Pictures\cpFactory_Conveyor.png
  5ce3da45-db07-42e7-a21c-a00fff4ed8f6|C:\Users\ggb\Documents\#PROJECTS\2016_06_29_Denmark\Pictures\071-050a_Bohren EA.jpg
  5ce3da45-db07-42e7-a21c-a00fff4ed8f6|C:\Users\ggb\Documents\#PROJECTS\2016_06_29_Denmark\Visu\RightArrow_Bold.png
  5ce3da45-db07-42e7-a21c-a00fff4ed8f6|C:\Users\ggb\Documents\#PROJECTS\2016_06_29_Denmark\Visu\German.gif
  5ce3da45-db07-42e7-a21c-a00fff4ed8f6|C:\Users\ggb\Documents\#PROJECTS\2016_06_29_Denmark\Visu\Parameters_1.png
  5ce3da45-db07-42e7-a21c-a00fff4ed8f6|C:\Users\ggb\Documents\#PROJECTS\2016_06_29_Denmark\Visu\Settings_1.png
  5ce3da45-db07-42e7-a21c-a00fff4ed8f6|C:\Users\ggb\Documents\#PROJECTS\2016_06_29_Denmark\Visu\Settings_1.png
  5ce3da45-db07-42e7-a21c-a00fff4ed8f6|C:\Users\ggb\Documents\#PROJECTS\2016_06_29_Denmark\Pictures\071-046b_Magazin.jpg
  5ce3da45-db07-42e7-a21c-a00fff4ed8f6|C:\Users\ggb\Documents\#PROJECTS\2016_06_29_Denmark\Pictures\cpFactory_Conveyor.png
  5ce3da45-db07-42e7-a21c-a00fff4ed8f6|C:\Users\ggb\Documents\#PROJECTS\2016_06_29_Denmark\Visu\Plus.png
  5ce3da45-db07-42e7-a21c-a00fff4ed8f6|C:\Users\ggb\Documents\#PROJECTS\2016_06_29_Denmark\Pictures\Kuka_Agilus.png